text list "SDC_EMS_FKT_INFO_REP": 0 'no maintenance text / No Repair Info'; 11 'drive: motor faulty / Drive: Drive 1 Defective'; 12 'drive: adjust scanner / Drive: Drive 2 Defective'; 13 'hoist: motor faulty / Hoist: Drive Defective'; 14 'hoist: adjust rope break switch / Tilt: Drive 1 Defective'; 15 'hoist: adjust reference height / Tilt: Drive 2 Defective'; 16 'hoist: adjust reference height initiator / Drive: Camera1 adjustment necessary'; 17 'spare / Drive: Camera2 adjustment necessary'; 18 'spare / Hoist: Camera2 adjustment necessary'; 19 'update software / Hoist: Ref-INI Camera1 adjustment necessary'; 20 'hardware changes / Tilt: Camera1 adjustment necessary'; 21 'spare / Tilt: Camera2 adjustment necessary'; 22 'update software / Tilt: Ref-INI Camera1 adjustment necessary'; 23 'spare / Repair info'; 24 'spare / Repair info'; 25 'spare / Repair info'; 26 'spare / Repair info'; 1 'PE-check / PE-Test'; 2 'brushs-check / Kohle-Test'; 3 'communication-check'

